(* Logix 5000 project; controller MV vendor 1 type 14 code 217 rev 31.11; software revision 31.00; part 12 of 53 *)
(* tags used below, declared in another part *)
   FVHRLTX02_IP : PlantItem;   // Effluent Tank Level Transmitter
   MC_B241 : INT[255];   // CH2 RN PMP Channel 2 return pum p drive flags
   MC_B243 : INT[255];   // CH2 ROUTE Channel 2 route requ est flags
   MC_CH2_CIP_BYPASS_Conditions : BOOL;
   MC_CH2_CIP_BYPASS_DrainConditions : BOOL;
   MC_CH2_DRAIN : PlantItem;   // CH2_DRAIN
   MC_CH2_LF1 : PlantItem;   // CH2_LF1
   MC_CH2_RR : PlantItem;   // CH2_RR
   MC_CH2_T125_2_ACC : DINT;
   MC_CIP_EFFTank_Start_Lvl_Ok : BOOL;
   MC_data_file_value_to_move : DINT;
   MC_N10 : INT[255];   // SETTINGS
   MC_N100 : INT[255];   // C1_PLC Channel 1 PLC data
   MC_N120 : INT[255];   // C2 PLC Channel 2 PLC data
   MC_N120_29_0_Storagebit : BOOL;
   MC_N122 : INT[255];   // CH2 PROG Channel 2 CIP progra m
   MC_N124 : INT[255];   // CH2 REPORT Channel 2 CIP report file
   MC_N80 : INT[255];   // SRV1_PLC Detergent tank 1 ser vice PLC data
   MC_N90 : INT[255];   // SV2_PLC Detergent tank 2 ser vice PLC data
   MC_T125 : TIMER[255];   // CH2 TIMERS Channel 2 timers
   MC_T4 : TIMER[255];   // TIMER
(* MC_Common, continued *)

ROUTINE MC_CH2_MCP_120   (* ladder *)
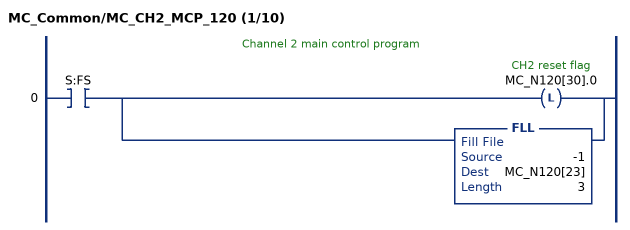
   // Channel 2 main control program
   0: XIC(S:FS)[OTL(MC_N120[30].0) ,FLL(-1,MC_N120[23],3) ];
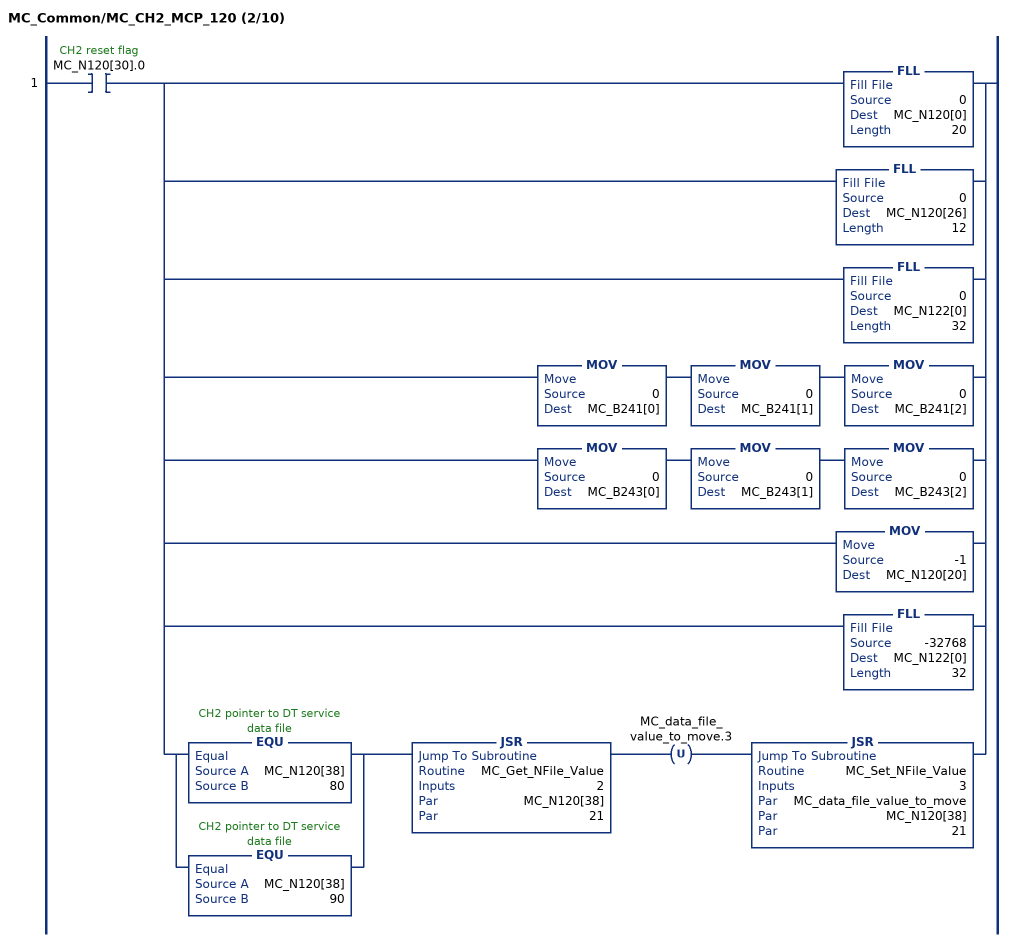
   1: XIC(MC_N120[30].0)[FLL(0,MC_N120[0],20) ,FLL(0,MC_N120[26],12) ,FLL(0,MC_N122[0],32) ,MOV(0,MC_B241[0]) MOV(0,MC_B241[1]) MOV(0,MC_B241[2]) ,MOV(0,MC_B243[0]) MOV(0,MC_B243[1]) MOV(0,MC_B243[2]) ,MOV(-1,MC_N120[20]) ,FLL(-32768,MC_N122[0],32) ,[EQU(MC_N120[38],80) ,EQU(MC_N120[38],90) ] JSR(MC_Get_NFile_Value,2,MC_N120[38],21) OTU(MC_data_file_value_to_move.3) JSR(MC_Set_NFile_Value,3,MC_data_file_value_to_move,MC_N120[38],21) ];
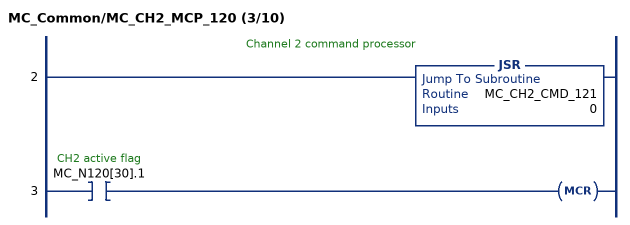
   // Channel 2 command processor
   2: JSR(MC_CH2_CMD_121,0);
   3: XIC(MC_N120[30].1)MCR();
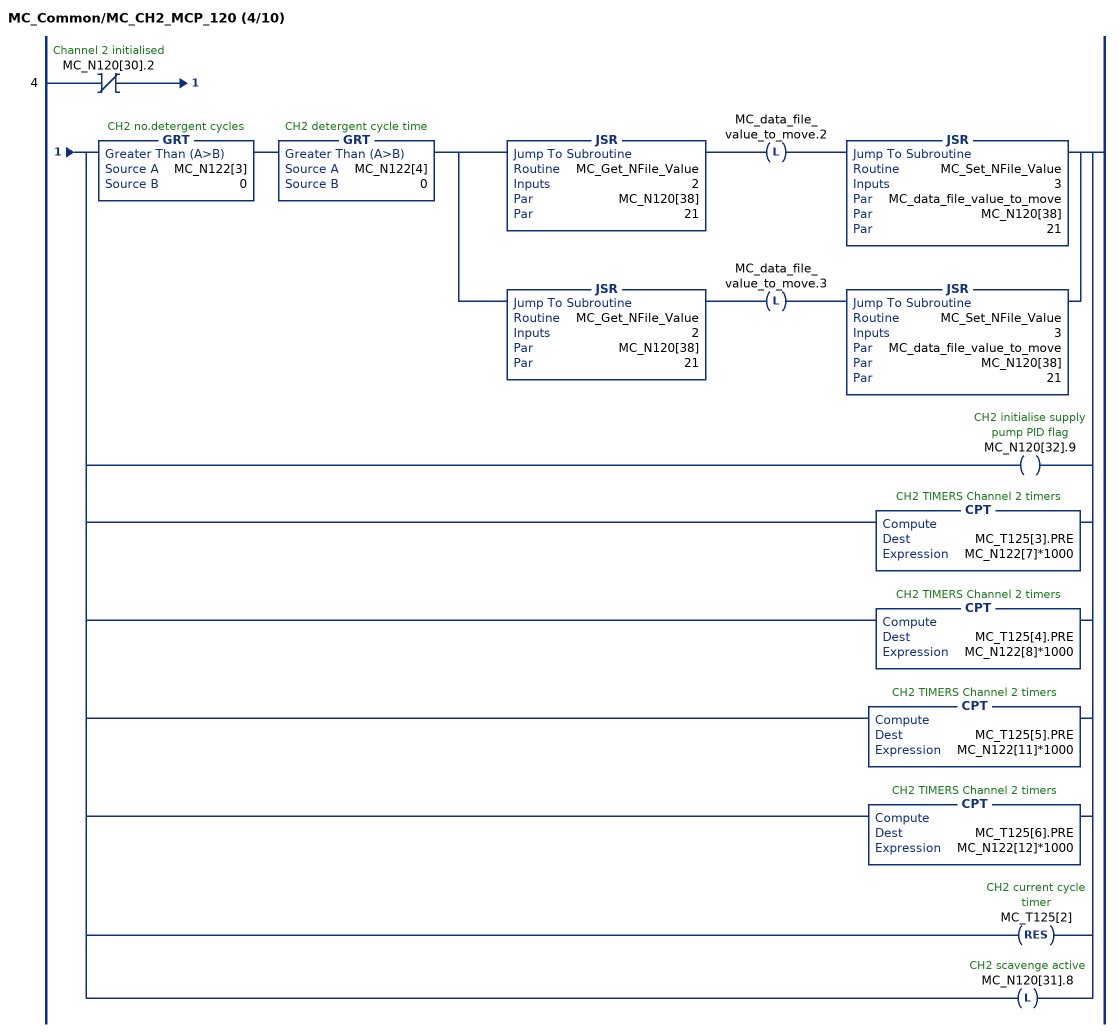
   4: XIO(MC_N120[30].2)[GRT(MC_N122[3],0) GRT(MC_N122[4],0) [JSR(MC_Get_NFile_Value,2,MC_N120[38],21) OTL(MC_data_file_value_to_move.2) JSR(MC_Set_NFile_Value,3,MC_data_file_value_to_move,MC_N120[38],21) ,JSR(MC_Get_NFile_Value,2,MC_N120[38],21) OTL(MC_data_file_value_to_move.3) JSR(MC_Set_NFile_Value,3,MC_data_file_value_to_move,MC_N120[38],21) ] ,OTE(MC_N120[32].9) ,[CPT(MC_T125[3].PRE,MC_N122[7]*1000) ,CPT(MC_T125[4].PRE,MC_N122[8]*1000) ,CPT(MC_T125[5].PRE,MC_N122[11]*1000) ,CPT(MC_T125[6].PRE,MC_N122[12]*1000) ,RES(MC_T125[2]) ,OTL(MC_N120[31].8) ] ];
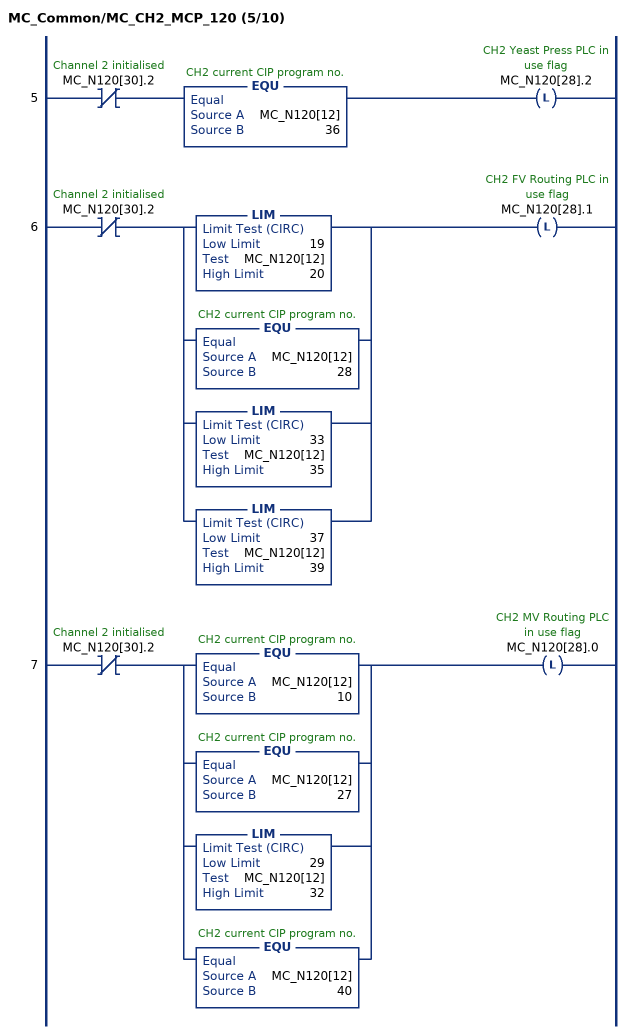
   5: XIO(MC_N120[30].2)EQU(MC_N120[12],36)OTL(MC_N120[28].2);
   6: XIO(MC_N120[30].2)[LIM(19,MC_N120[12],20) ,EQU(MC_N120[12],28) ,LIM(33,MC_N120[12],35) ,LIM(37,MC_N120[12],39) ]OTL(MC_N120[28].1);
   7: XIO(MC_N120[30].2)[EQU(MC_N120[12],10) ,EQU(MC_N120[12],27) ,LIM(29,MC_N120[12],32) ,EQU(MC_N120[12],40) ]OTL(MC_N120[28].0);
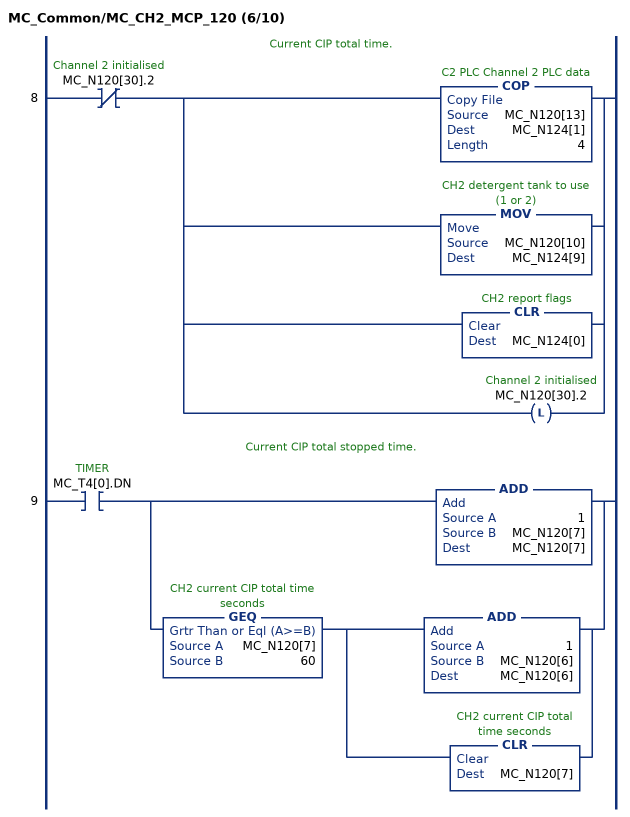
   // Current CIP total time.
   8: XIO(MC_N120[30].2)[COP(MC_N120[13],MC_N124[1],4) ,MOV(MC_N120[10],MC_N124[9]) ,CLR(MC_N124[0]) ,OTL(MC_N120[30].2) ];
   // Current CIP total stopped time.
   9: XIC(MC_T4[0].DN)[ADD(1,MC_N120[7],MC_N120[7]) ,GEQ(MC_N120[7],60) [ADD(1,MC_N120[6],MC_N120[6]) ,CLR(MC_N120[7]) ] ];
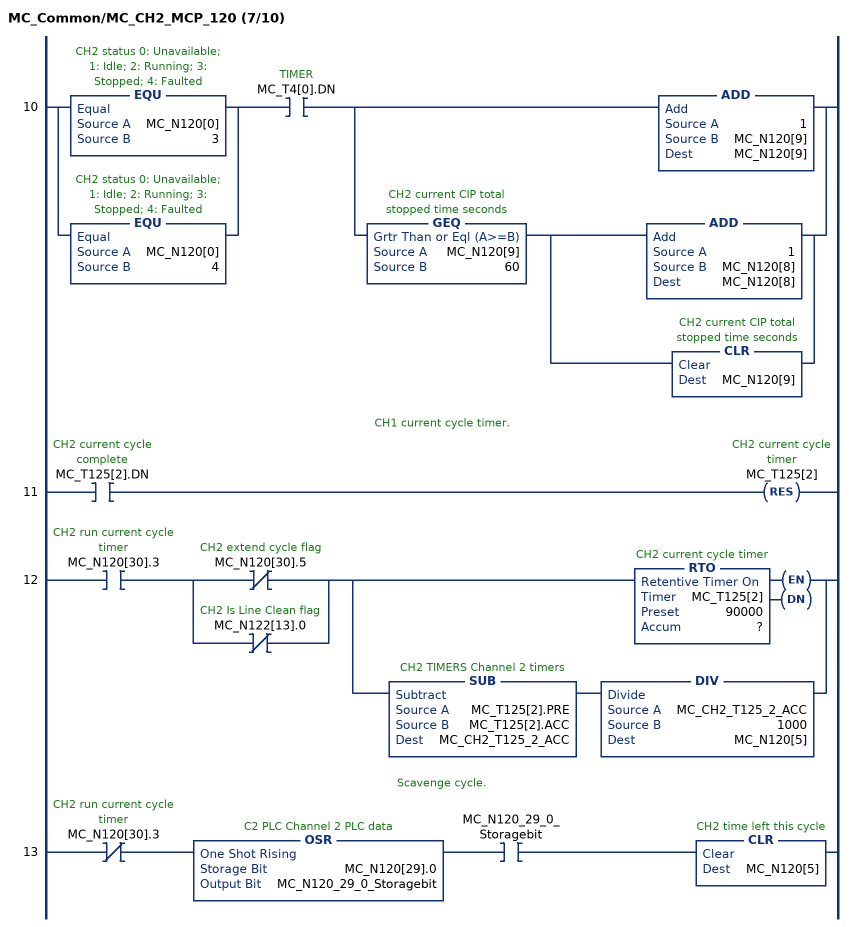
   10: [EQU(MC_N120[0],3) ,EQU(MC_N120[0],4) ]XIC(MC_T4[0].DN)[ADD(1,MC_N120[9],MC_N120[9]) ,GEQ(MC_N120[9],60) [ADD(1,MC_N120[8],MC_N120[8]) ,CLR(MC_N120[9]) ] ];
   // CH1 current cycle timer.
   11: XIC(MC_T125[2].DN)RES(MC_T125[2]);
   12: XIC(MC_N120[30].3)[XIO(MC_N120[30].5) ,XIO(MC_N122[13].0) ][RTO(MC_T125[2],?,?) ,SUB(MC_T125[2].PRE,MC_T125[2].ACC,MC_CH2_T125_2_ACC) DIV(MC_CH2_T125_2_ACC,1000,MC_N120[5]) ];
   // Scavenge cycle.
   13: XIO(MC_N120[30].3)OSR(MC_N120[29].0,MC_N120_29_0_Storagebit)XIC(MC_N120_29_0_Storagebit)CLR(MC_N120[5]);
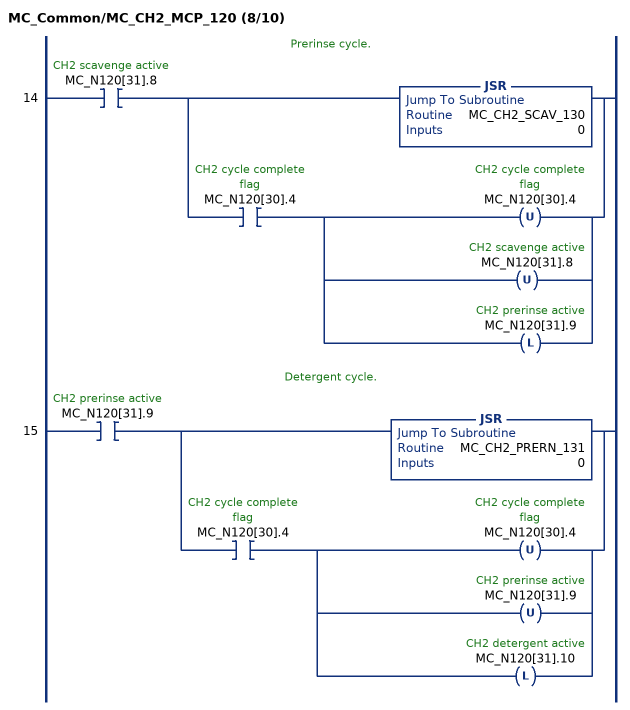
   // Prerinse cycle.
   14: XIC(MC_N120[31].8)[JSR(MC_CH2_SCAV_130,0) ,XIC(MC_N120[30].4) [OTU(MC_N120[30].4) ,OTU(MC_N120[31].8) ,OTL(MC_N120[31].9) ] ];
   // Detergent cycle.
   15: XIC(MC_N120[31].9)[JSR(MC_CH2_PRERN_131,0) ,XIC(MC_N120[30].4) [OTU(MC_N120[30].4) ,OTU(MC_N120[31].9) ,OTL(MC_N120[31].10) ] ];
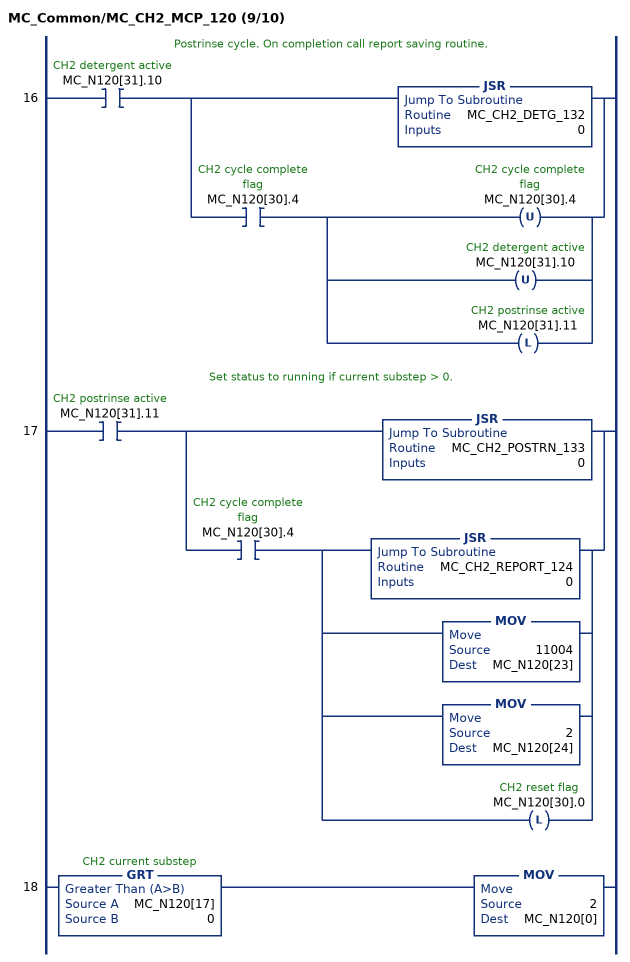
   // Postrinse cycle. On completion call report saving routine.
   16: XIC(MC_N120[31].10)[JSR(MC_CH2_DETG_132,0) ,XIC(MC_N120[30].4) [OTU(MC_N120[30].4) ,OTU(MC_N120[31].10) ,OTL(MC_N120[31].11) ] ];
   // Set status to running if current substep > 0.
   17: XIC(MC_N120[31].11)[JSR(MC_CH2_POSTRN_133,0) ,XIC(MC_N120[30].4) [JSR(MC_CH2_REPORT_124,0) ,MOV(11004,MC_N120[23]) ,MOV(2,MC_N120[24]) ,OTL(MC_N120[30].0) ] ];
   18: GRT(MC_N120[17],0)MOV(2,MC_N120[0]);
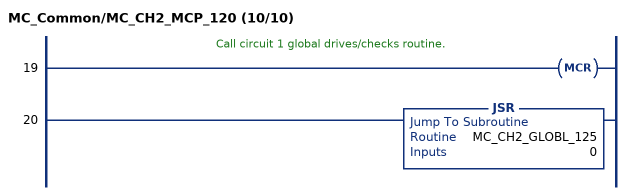
   // Call circuit 1 global drives/checks routine.
   19: MCR();
   20: JSR(MC_CH2_GLOBL_125,0);
END_ROUTINE

ROUTINE MC_CH2_POSTRN_133   (* ladder *)
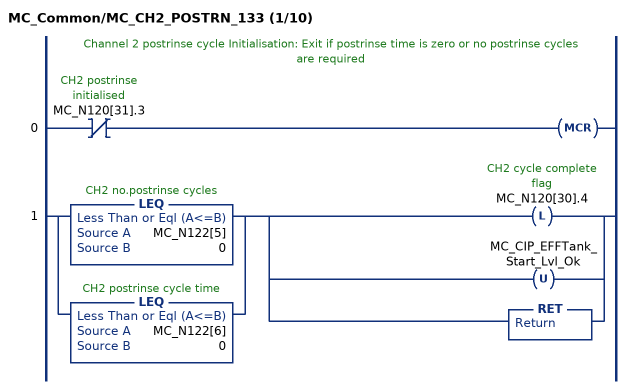
   // Channel 2 postrinse cycle Initialisation: Exit if postrinse time is zero or no postrinse cycles are required
   0: XIO(MC_N120[31].3)MCR();
   1: [LEQ(MC_N122[5],0) ,LEQ(MC_N122[6],0) ][OTL(MC_N120[30].4) ,OTU(MC_CIP_EFFTank_Start_Lvl_Ok) ,RET() ];
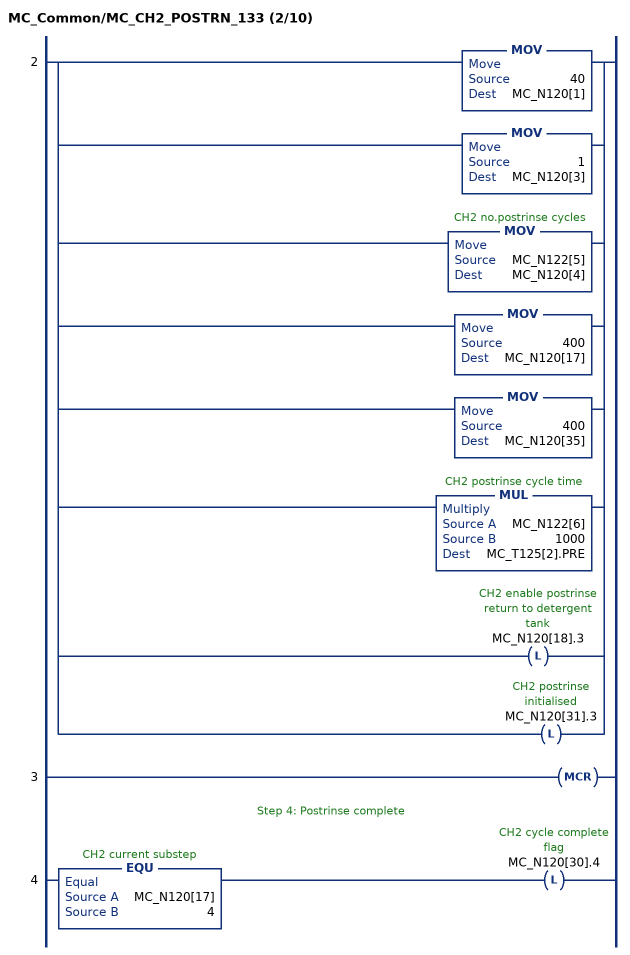
   2: [MOV(40,MC_N120[1]) ,MOV(1,MC_N120[3]) ,MOV(MC_N122[5],MC_N120[4]) ,MOV(400,MC_N120[17]) ,MOV(400,MC_N120[35]) ,MUL(MC_N122[6],1000,MC_T125[2].PRE) ,OTL(MC_N120[18].3) ,OTL(MC_N120[31].3) ];
   3: MCR();
   // Step 4: Postrinse complete
   4: EQU(MC_N120[17],4)OTL(MC_N120[30].4);
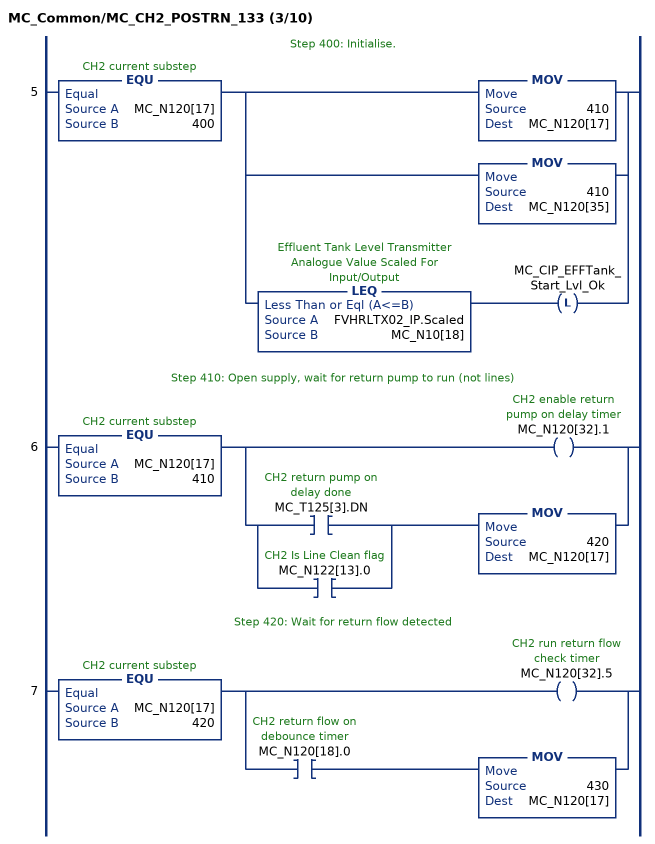
   // Step 400: Initialise.
   5: EQU(MC_N120[17],400)[MOV(410,MC_N120[17]) ,MOV(410,MC_N120[35]) ,LEQ(FVHRLTX02_IP.Scaled,MC_N10[18]) OTL(MC_CIP_EFFTank_Start_Lvl_Ok) ];
   // Step 410: Open supply, wait for return pump to run (not lines)
   6: EQU(MC_N120[17],410)[OTE(MC_N120[32].1) ,[XIC(MC_T125[3].DN) ,XIC(MC_N122[13].0) ] MOV(420,MC_N120[17]) ];
   // Step 420: Wait for return flow detected
   7: EQU(MC_N120[17],420)[OTE(MC_N120[32].5) ,XIC(MC_N120[18].0) MOV(430,MC_N120[17]) ];
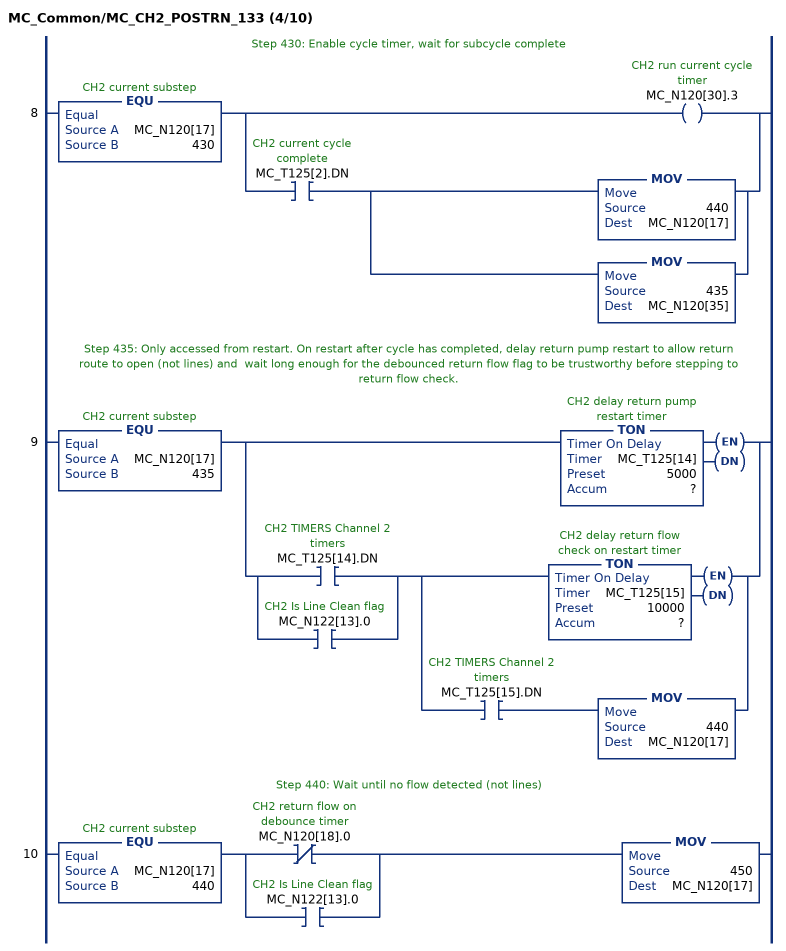
   // Step 430: Enable cycle timer, wait for subcycle complete
   8: EQU(MC_N120[17],430)[OTE(MC_N120[30].3) ,XIC(MC_T125[2].DN) [MOV(440,MC_N120[17]) ,MOV(435,MC_N120[35]) ] ];
   // Step 435: Only accessed from restart. On restart after cycle has completed, delay return pump restart to allow return route to open (not lines) and  wait long enough for the debounced return flow flag to be trustworthy before stepping to return flow check.
   9: EQU(MC_N120[17],435)[TON(MC_T125[14],?,?) ,[XIC(MC_T125[14].DN) ,XIC(MC_N122[13].0) ] [TON(MC_T125[15],?,?) ,XIC(MC_T125[15].DN) MOV(440,MC_N120[17]) ] ];
   // Step 440: Wait until no flow detected (not lines)
   10: EQU(MC_N120[17],440)[XIO(MC_N120[18].0) ,XIC(MC_N122[13].0) ]MOV(450,MC_N120[17]);
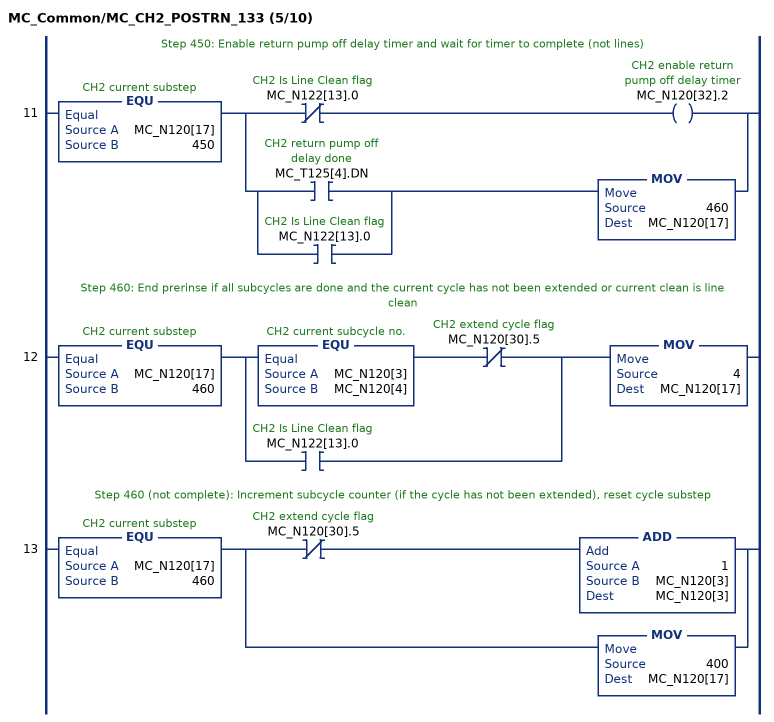
   // Step 450: Enable return pump off delay timer and wait for timer to complete (not lines)
   11: EQU(MC_N120[17],450)[XIO(MC_N122[13].0) OTE(MC_N120[32].2) ,[XIC(MC_T125[4].DN) ,XIC(MC_N122[13].0) ] MOV(460,MC_N120[17]) ];
   // Step 460: End prerinse if all subcycles are done and the current cycle has not been extended or current clean is line clean
   12: EQU(MC_N120[17],460)[EQU(MC_N120[3],MC_N120[4]) XIO(MC_N120[30].5) ,XIC(MC_N122[13].0) ]MOV(4,MC_N120[17]);
   // Step 460 (not complete): Increment subcycle counter (if the cycle has not been extended), reset cycle substep
   13: EQU(MC_N120[17],460)[XIO(MC_N120[30].5) ADD(1,MC_N120[3],MC_N120[3]) ,MOV(400,MC_N120[17]) ];
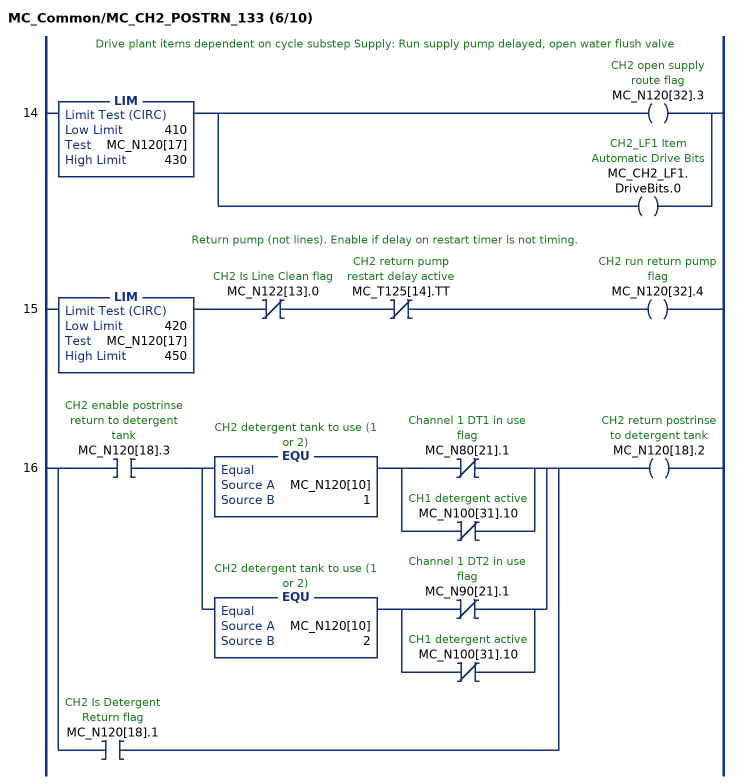
   // Drive plant items dependent on cycle substep Supply: Run supply pump delayed, open water flush valve
   14: LIM(410,MC_N120[17],430)[OTE(MC_N120[32].3) ,OTE(MC_CH2_LF1.DriveBits.0) ];
   // Return pump (not lines). Enable if delay on restart timer is not timing.
   15: LIM(420,MC_N120[17],450)XIO(MC_N122[13].0)XIO(MC_T125[14].TT)OTE(MC_N120[32].4);
   16: [XIC(MC_N120[18].3) [EQU(MC_N120[10],1) [XIO(MC_N80[21].1) ,XIO(MC_N100[31].10) ] ,EQU(MC_N120[10],2) [XIO(MC_N90[21].1) ,XIO(MC_N100[31].10) ] ] ,XIC(MC_N120[18].1) ]OTE(MC_N120[18].2);
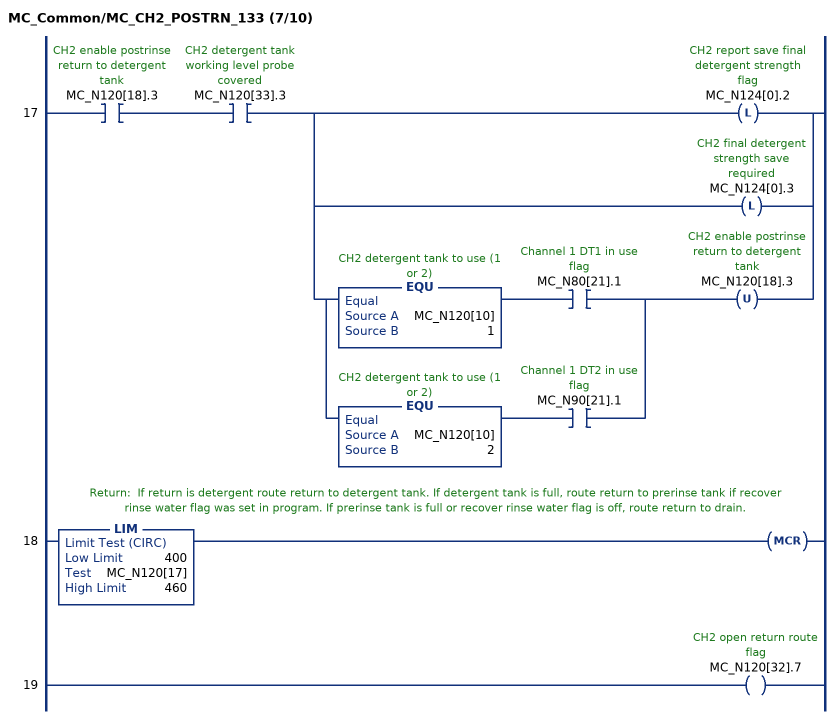
   17: XIC(MC_N120[18].3)XIC(MC_N120[33].3)[OTL(MC_N124[0].2) ,OTL(MC_N124[0].3) ,[EQU(MC_N120[10],1) XIC(MC_N80[21].1) ,EQU(MC_N120[10],2) XIC(MC_N90[21].1) ] OTU(MC_N120[18].3) ];
   // Return:  If return is detergent route return to detergent tank. If detergent tank is full, route return to prerinse tank if recover rinse water flag was set in program. If prerinse tank is full or recover rinse water flag is off, route return to drain.
   18: LIM(400,MC_N120[17],460)MCR();
   19: OTE(MC_N120[32].7);
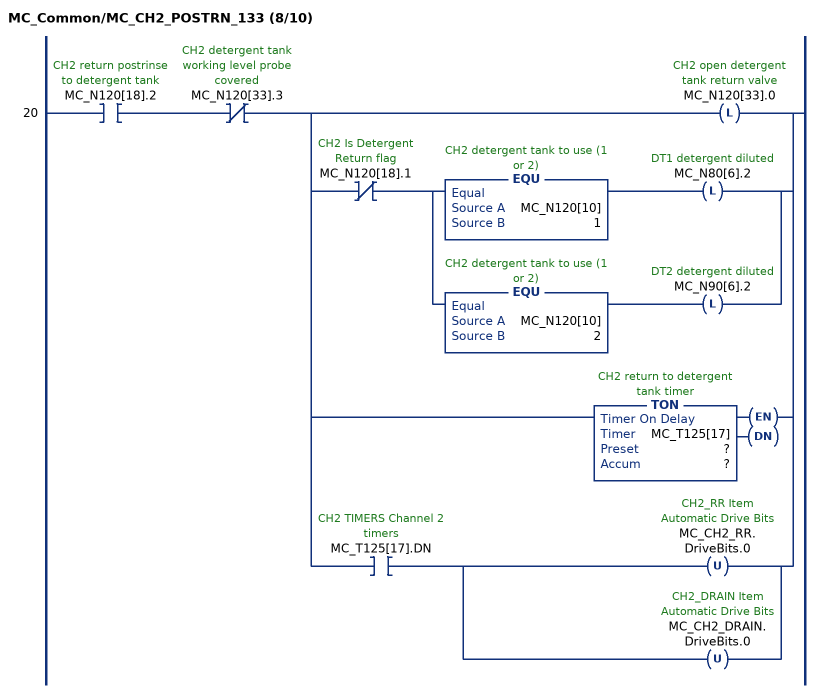
   20: XIC(MC_N120[18].2)XIO(MC_N120[33].3)[OTL(MC_N120[33].0) ,XIO(MC_N120[18].1) [EQU(MC_N120[10],1) OTL(MC_N80[6].2) ,EQU(MC_N120[10],2) OTL(MC_N90[6].2) ] ,TON(MC_T125[17],?,?) ,XIC(MC_T125[17].DN) [OTU(MC_CH2_RR.DriveBits.0) ,OTU(MC_CH2_DRAIN.DriveBits.0) ] ];
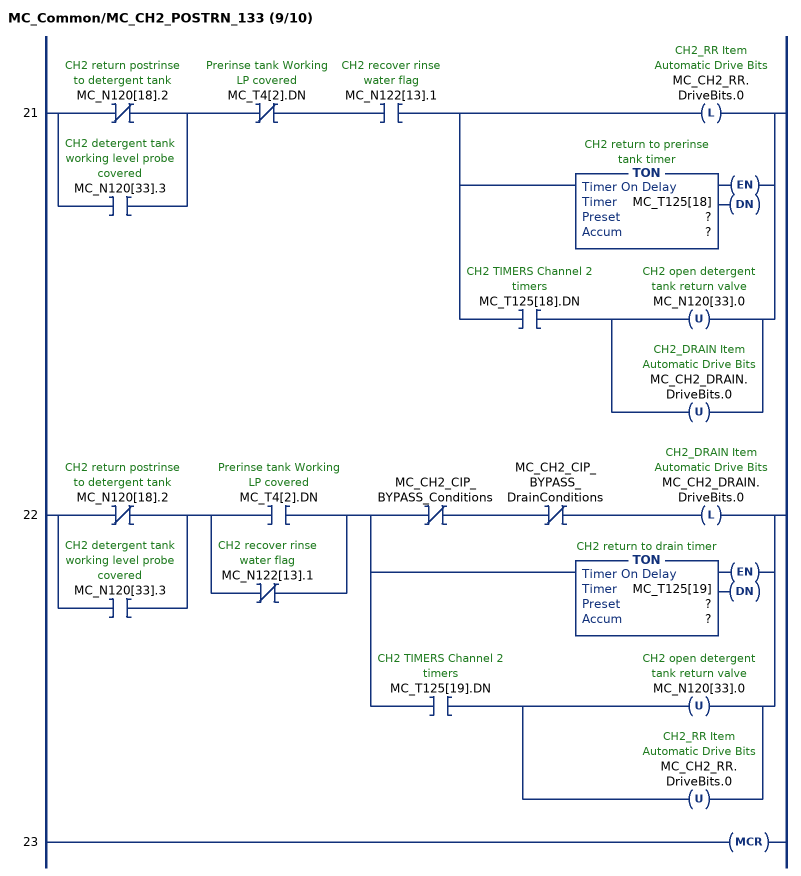
   21: [XIO(MC_N120[18].2) ,XIC(MC_N120[33].3) ]XIO(MC_T4[2].DN)XIC(MC_N122[13].1)[OTL(MC_CH2_RR.DriveBits.0) ,TON(MC_T125[18],?,?) ,XIC(MC_T125[18].DN) [OTU(MC_N120[33].0) ,OTU(MC_CH2_DRAIN.DriveBits.0) ] ];
   22: [XIO(MC_N120[18].2) ,XIC(MC_N120[33].3) ][XIC(MC_T4[2].DN) ,XIO(MC_N122[13].1) ][XIO(MC_CH2_CIP_BYPASS_Conditions) XIO(MC_CH2_CIP_BYPASS_DrainConditions) OTL(MC_CH2_DRAIN.DriveBits.0) ,TON(MC_T125[19],?,?) ,XIC(MC_T125[19].DN) [OTU(MC_N120[33].0) ,OTU(MC_CH2_RR.DriveBits.0) ] ];
   23: MCR();
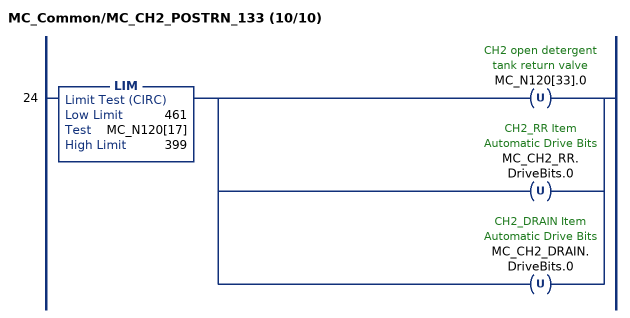
   24: LIM(461,MC_N120[17],399)[OTU(MC_N120[33].0) ,OTU(MC_CH2_RR.DriveBits.0) ,OTU(MC_CH2_DRAIN.DriveBits.0) ];
END_ROUTINE
